VERSION : 0.1
   VAR_INPUT
      IN1 : DInt;
      IN2 : DInt;
      IN3 : DInt;
      IN4 : DInt;
      IN5 : DInt;
      IN6 : DInt;
      IN7 : DInt;
   END_VAR
   VAR_OUTPUT
      Out : Real;
   END_VAR
BEGIN

REGION Network 2 (SCL)
   #Out := (DINT_TO_REAL(#IN1 + #IN2 + #IN3) - DINT_TO_REAL(#IN4 + #IN5 + #IN6)) / #IN7;
END_REGION
END_FUNCTION_BLOCK

FUNCTION_BLOCK "PGC Flush"   // FB517, LAD
{ S7_Optimized_Access := 'TRUE' }
VERSION : 0.1
   VAR_INPUT
      Activate : Bool;
      Override : Bool;
      "PGC Purge Duration" : Time := T#60m;
      "Temperature Setpoint" : Real := 50.0;
      Temperature : Real;
      "PGC Stop Delay" : Time := T#10m;
      "PGC Stoped" : Bool;
      "CAB Started" : Bool;
      "CAB after Start Delay" : Time := T#60s;
      "CAB RPM Cmd" : Real := 400.0;
      "IGG Mode" : Int;   // 1 = Auto, 2 = Man, 3 = FatAuto, 4 = FatMan
      "IGG Stoped" : Bool;
      Alarm : Bool;
      "CV405 Opened" : Real;
      "CV403 Opened" : Real;
      "CV401 Opened" : Bool;
      "CV441 Closed" : Bool;
      "CV431 Opened" : Bool;
   END_VAR
   VAR_OUTPUT
      "CV405 Open" : Bool;
      "CV403 Open" : Bool;
      "CV401 Open" : Bool;
      "CV441 Close" : Bool;
      "CV431 Open" : Bool;
      "CAB Start" : Bool;
      "CAB RPM Ctrl" : Real;
      "CV403 Modulate" : Bool;
      Running : Bool;
      "Stop PGC" : Bool;
      Done : Bool;
   END_VAR
   VAR
      "CAB earlier Stop Aux" : Time;
      "PGC Stop Delay TON" : TON_TIME;
      "Sequence Max Time TON" : TON_TIME;
      "CAB after Start Delay TON" : TON_TIME;
      "Flip Flop_Override" : "Flip Flop";
      "CAB earlier STOP" : TON_TIME;
      "Valve to origin Delay" : TOF_TIME;
      "Valve Opened Delay" : TOF_TIME;
      "PGC Stop Puls" : TP_TIME;
      "Modulate Delay" : TON_TIME;
      "CAB after Start Delay Aux" : Bool;
   END_VAR
BEGIN

REGION Network 1
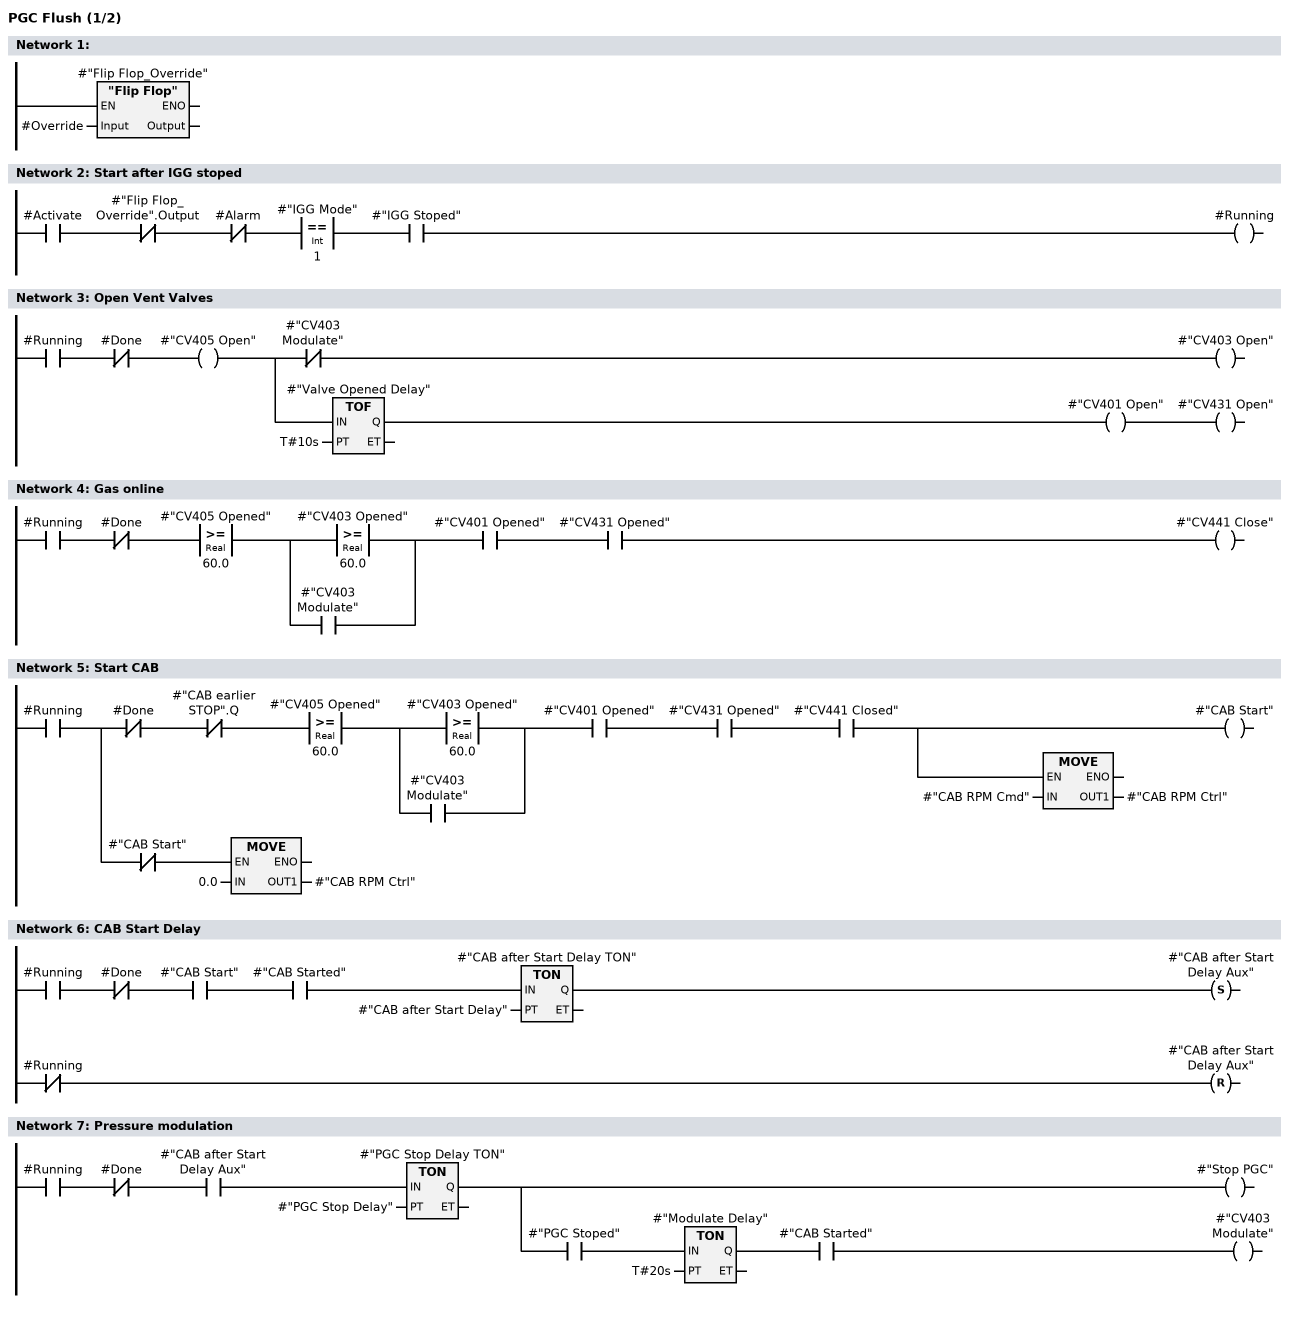
   RUNG wire#powerrail
      #"Flip Flop_Override"(Input := #Override, Output =>)
   END_RUNG
   // the same network as SCL:
   #"Flip Flop_Override"(Input := #Override);   // "Flip Flop"
END_REGION

REGION Network 2: Start after IGG stoped
   RUNG wire#powerrail
      Contact( #Activate )
      I_Contact( #"Flip Flop_Override".Output )
      I_Contact( #Alarm )
      { S7_Templates := "SrcType := Int" } EQ_Contact(in1 := #"IGG Mode", in2 := 1)
      Contact( #"IGG Stoped" )
      Coil( #Running )
   END_RUNG
   // the same network as SCL:
   #Running := #Activate AND NOT #"Flip Flop_Override".Output AND NOT #Alarm AND (#"IGG Mode" = 1) AND #"IGG Stoped";
END_REGION

REGION Network 3: Open Vent Valves
   #"CV405 Open" := #Running AND NOT #Done;
   #"CV403 Open" := #"CV405 Open" AND NOT #"CV403 Modulate";
   #"Valve Opened Delay"(IN := #"CV405 Open", PT := T#10s);   // TOF
   #"CV401 Open" := #"Valve Opened Delay".Q;
   #"CV431 Open" := #"Valve Opened Delay".Q;
END_REGION

REGION Network 4: Gas online
   RUNG wire#powerrail
      Contact( #Running )
      I_Contact( #Done )
      { S7_Templates := "SrcType := Real" } GE_Contact(in1 := #"CV405 Opened", in2 := 60.0)
      wire#w1
      { S7_Templates := "SrcType := Real" } GE_Contact(in1 := #"CV403 Opened", in2 := 60.0)
      wire#w2
      Contact( #"CV401 Opened" )
      Contact( #"CV431 Opened" )
      Coil( #"CV441 Close" )
   END_RUNG
   RUNG wire#w1
      Contact( #"CV403 Modulate" )
   END_RUNG wire#w2
   // the same network as SCL:
   #"CV441 Close" := #Running AND NOT #Done AND (#"CV405 Opened" >= 60.0) AND ((#"CV403 Opened" >= 60.0) OR #"CV403 Modulate") AND #"CV401 Opened" AND #"CV431 Opened";
END_REGION

REGION Network 5: Start CAB
   RUNG wire#powerrail
      Contact( #Running )
      wire#w1
      I_Contact( #Done )
      I_Contact( #"CAB earlier STOP".Q )
      { S7_Templates := "SrcType := Real" } GE_Contact(in1 := #"CV405 Opened", in2 := 60.0)
      wire#w2
      { S7_Templates := "SrcType := Real" } GE_Contact(in1 := #"CV403 Opened", in2 := 60.0)
      wire#w3
      Contact( #"CV401 Opened" )
      Contact( #"CV431 Opened" )
      Contact( #"CV441 Closed" )
      wire#w4
      Coil( #"CAB Start" )
   END_RUNG
   RUNG wire#w2
      Contact( #"CV403 Modulate" )
   END_RUNG wire#w3
   RUNG wire#w4
      Move(in := #"CAB RPM Cmd", out1 => #"CAB RPM Ctrl")
   END_RUNG
   RUNG wire#w1
      I_Contact( #"CAB Start" )
      Move(in := 0.0, out1 => #"CAB RPM Ctrl")
   END_RUNG
   // the same network as SCL:
   #"CAB Start" := #Running AND NOT #Done AND NOT #"CAB earlier STOP".Q AND (#"CV405 Opened" >= 60.0) AND ((#"CV403 Opened" >= 60.0) OR #"CV403 Modulate") AND #"CV401 Opened" AND #"CV431 Opened" AND #"CV441 Closed";
   IF #"CAB Start" THEN #"CAB RPM Ctrl" := #"CAB RPM Cmd"; END_IF;
   IF #Running AND NOT #"CAB Start" THEN #"CAB RPM Ctrl" := 0.0; END_IF;
END_REGION

REGION Network 6: CAB Start Delay
   #"CAB after Start Delay TON"(IN := #Running AND NOT #Done AND #"CAB Start" AND #"CAB Started",   // TON
                           PT := #"CAB after Start Delay");
   IF #"CAB after Start Delay TON".Q THEN #"CAB after Start Delay Aux" := TRUE; END_IF;
   IF NOT #Running THEN #"CAB after Start Delay Aux" := FALSE; END_IF;
END_REGION

REGION Network 7: Pressure modulation
   #"PGC Stop Delay TON"(IN := #Running AND NOT #Done AND #"CAB after Start Delay Aux", PT := #"PGC Stop Delay");   // TON
   #"Stop PGC" := #"PGC Stop Delay TON".Q;
   #"Modulate Delay"(IN := #"PGC Stop Delay TON".Q AND #"PGC Stoped", PT := T#20s);   // TON
   #"CV403 Modulate" := #"Modulate Delay".Q AND #"CAB Started";
END_REGION

REGION Network 8: Sequence max time
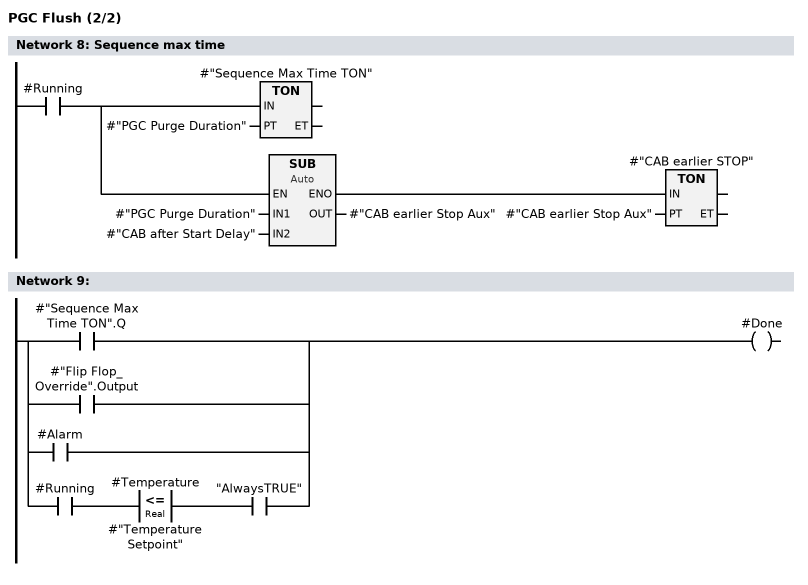
   #"Sequence Max Time TON"(IN := #Running, PT := #"PGC Purge Duration");   // TON
   IF #Running THEN #"CAB earlier Stop Aux" := #"PGC Purge Duration" - #"CAB after Start Delay"; END_IF;
   #"CAB earlier STOP"(IN := #Running, PT := #"CAB earlier Stop Aux");   // TON
END_REGION

REGION Network 9
   RUNG wire#powerrail
      Contact( #"Sequence Max Time TON".Q )
      wire#w1
      Coil( #Done )
   END_RUNG
   RUNG wire#powerrail
      Contact( #"Flip Flop_Override".Output )
   END_RUNG wire#w1
   RUNG wire#powerrail
      Contact( #Alarm )
   END_RUNG wire#w1
   RUNG wire#powerrail
      Contact( #Running )
      { S7_Templates := "SrcType := Real" } LE_Contact(in1 := #Temperature, in2 := #"Temperature Setpoint")
      Contact( "AlwaysTRUE" )
   END_RUNG wire#w1
   // the same network as SCL:
   #Done := #"Sequence Max Time TON".Q OR #"Flip Flop_Override".Output OR #Alarm OR (#Running AND (#Temperature <= #"Temperature Setpoint") AND "AlwaysTRUE");
END_REGION
END_FUNCTION_BLOCK

FUNCTION_BLOCK "RAMP"   // FB518, LAD
{ S7_Optimized_Access := 'TRUE' }
VERSION : 0.1
   VAR_INPUT
      Start : Bool;
      "Time span" : Time;
      "Minimum Value" : Real;
      "Maximum Value" : Real;
   END_VAR
   VAR_OUTPUT
      Value : Real;
      "Ramp Done" : Bool;
   END_VAR
   VAR
      "RUN Time" : TON_TIME;
      "RUN Time Aux" : Real;
      "Time span Aux" : Real;
      "Maximum Value M" : Real;
   END_VAR
BEGIN

REGION Network 1
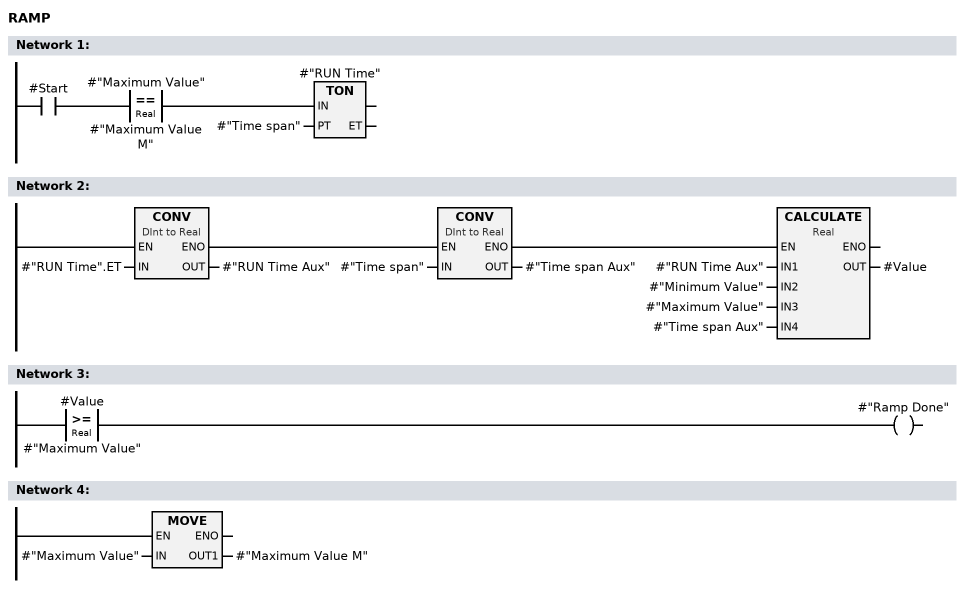
   #"RUN Time"(IN := #Start AND (#"Maximum Value" = #"Maximum Value M"), PT := #"Time span");   // TON
END_REGION

REGION Network 2
   RUNG wire#powerrail
      { S7_Templates := "[SrcType := DInt, DestType := Real]" } Convert(in := #"RUN Time".ET, out => #"RUN Time Aux")
      { S7_Templates := "[SrcType := DInt, DestType := Real]" } Convert(in := #"Time span", out => #"Time span Aux")
      { S7_Templates := "SrcType := Real"; S7_Expression := "((IN1*(IN3-IN2))/IN4)+IN2" } Calculate(in1 := #"RUN Time Aux", in2 := #"Minimum Value", in3 := #"Maximum Value", in4 := #"Time span Aux", out => #Value)
   END_RUNG
   // the same network as SCL:
   #"RUN Time Aux" := DINT_TO_REAL(#"RUN Time".ET);
   #"Time span Aux" := DINT_TO_REAL(#"Time span");
   #Value := ((#"RUN Time Aux"*(#"Maximum Value"-#"Minimum Value"))/#"Time span Aux")+#"Minimum Value";
END_REGION

REGION Network 3
   RUNG wire#powerrail
      { S7_Templates := "SrcType := Real" } GE_Contact(in1 := #Value, in2 := #"Maximum Value")
      Coil( #"Ramp Done" )
   END_RUNG
   // the same network as SCL:
   #"Ramp Done" := #Value >= #"Maximum Value";
END_REGION

REGION Network 4
   RUNG wire#powerrail
      Move(in := #"Maximum Value", out1 => #"Maximum Value M")
   END_RUNG
   // the same network as SCL:
   #"Maximum Value M" := #"Maximum Value";
END_REGION
END_FUNCTION_BLOCK

FUNCTION_BLOCK "Choose Real"   // FB519, LAD
{ S7_Optimized_Access := 'TRUE' }
VERSION : 0.1
   VAR_INPUT
      Choose : Bool;
      "Option 1" : Real;
      "Option 2" : Real;
   END_VAR
   VAR_OUTPUT
      Output : Real;
   END_VAR
   VAR
      True : Bool;
      False : Bool;
      "Option 1 M" : Real;
      "Option 2 M" : Real;
      "Choose Internal" : Bool;
      "Puls Aux" : Struct
         "Puls Aux 1" : Bool;
         "Puls Aux 2" : Bool;
         "Puls Aux 3" : Bool;
         "Puls Aux 4" : Bool;
         "Puls Aux 5" : Bool;
         "Puls Aux 6" : Bool;
      END_STRUCT;
      "TP P CHOOSE1" : TP_TIME;
      "TP N CHOOSE2" : TP_TIME;
      "TP N CHOOSE1" : TP_TIME;
      "TP P CHOOSE2" : TP_TIME;
      R_TRIG_Instance : R_TRIG;
      Puls : TP_TIME;
   END_VAR
   VAR_TEMP   // added for the SCL form of the ladder/FBD networks
      _w1 : Bool;
      _w2 : Bool;
      _w3 : Bool;
      _w4 : Bool;
      _w5 : Bool;
   END_VAR
BEGIN

REGION Network 1: False/True
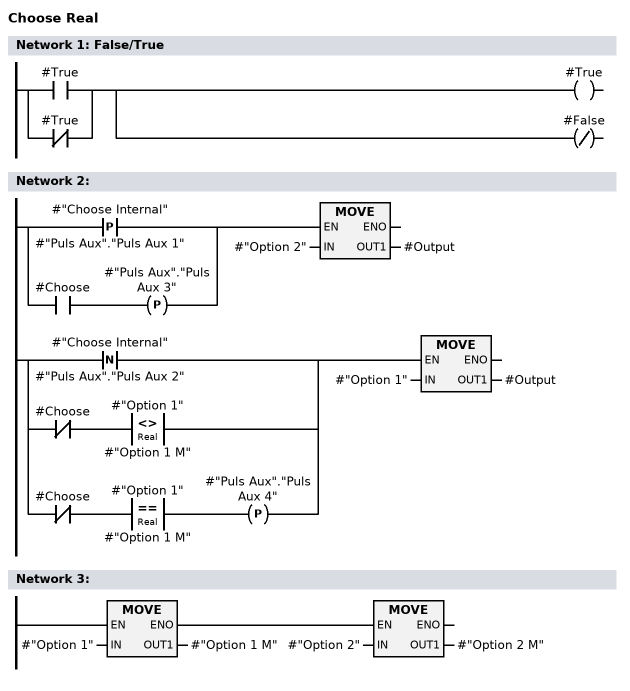
   RUNG wire#powerrail
      Contact( #True )
      wire#w1
      Coil( #True )
   END_RUNG
   RUNG wire#powerrail
      I_Contact( #True )
   END_RUNG wire#w1
   RUNG wire#w1
      I_Coil( #False )
   END_RUNG
   // the same network as SCL:
   #True := #True OR NOT #True;
   #False := NOT #True;
END_REGION

REGION Network 2
   RUNG wire#powerrail
      P_Contact(operand := #"Choose Internal", bit := #"Puls Aux"."Puls Aux 1")
      wire#w1
      Move(in := #"Option 2", out1 => #Output)
   END_RUNG
   RUNG wire#powerrail
      Contact( #Choose )
      P_Trig( #"Puls Aux"."Puls Aux 3" )
   END_RUNG wire#w1
   RUNG wire#powerrail
      N_Contact(operand := #"Choose Internal", bit := #"Puls Aux"."Puls Aux 2")
      wire#w2
      Move(in := #"Option 1", out1 => #Output)
   END_RUNG
   RUNG wire#powerrail
      I_Contact( #Choose )
      { S7_Templates := "SrcType := Real" } NE_Contact(in1 := #"Option 1", in2 := #"Option 1 M")
   END_RUNG wire#w2
   RUNG wire#powerrail
      I_Contact( #Choose )
      { S7_Templates := "SrcType := Real" } EQ_Contact(in1 := #"Option 1", in2 := #"Option 1 M")
      P_Trig( #"Puls Aux"."Puls Aux 4" )
   END_RUNG wire#w2
   // the same network as SCL:
   #_w1 := #"Choose Internal" AND NOT #"Puls Aux"."Puls Aux 1";   // rising edge of #"Choose Internal"
   #"Puls Aux"."Puls Aux 1" := #"Choose Internal";
   #_w2 := #Choose AND NOT #"Puls Aux"."Puls Aux 3";   // rising edge
   #"Puls Aux"."Puls Aux 3" := #Choose;
   IF #_w1 OR #_w2 THEN #Output := #"Option 2"; END_IF;
   #_w3 := NOT #"Choose Internal" AND #"Puls Aux"."Puls Aux 2";   // falling edge of #"Choose Internal"
   #"Puls Aux"."Puls Aux 2" := #"Choose Internal";
   #_w4 := NOT #Choose AND (#"Option 1" = #"Option 1 M");
   #_w5 := #_w4 AND NOT #"Puls Aux"."Puls Aux 4";   // rising edge
   #"Puls Aux"."Puls Aux 4" := #_w4;
   IF #_w3 OR (NOT #Choose AND (#"Option 1" <> #"Option 1 M")) OR #_w5 THEN #Output := #"Option 1"; END_IF;
END_REGION

REGION Network 3
   RUNG wire#powerrail
      Move(in := #"Option 1", out1 => #"Option 1 M")
      Move(in := #"Option 2", out1 => #"Option 2 M")
   END_RUNG
   // the same network as SCL:
   #"Option 1 M" := #"Option 1";
   #"Option 2 M" := #"Option 2";
END_REGION
END_FUNCTION_BLOCK

FUNCTION "Bool to Word" : Void   // FC202, FBD
{ S7_Optimized_Access := 'FALSE' }
VERSION : 0.1
// Die Funktion gruppiert 16 Variablen vom Datentyp "Bool" zu einer Variablen vom Datentyp "Word".
// *******************************************************************************
// The function groups 16 variables with type of data "Bool" to a variable with type of data "Word".
   VAR_INPUT
      Bit0 : Bool;
      Bit1 : Bool;
      Bit2 : Bool;
      Bit3 : Bool;
      Bit4 : Bool;
      Bit5 : Bool;
      Bit6 : Bool;
      Bit7 : Bool;
      Bit8 : Bool;
      Bit9 : Bool;
      Bit10 : Bool;
      Bit11 : Bool;
      Bit12 : Bool;
      Bit13 : Bool;
      Bit14 : Bool;
      Bit15 : Bool;
   END_VAR
   VAR_OUTPUT
      "Word" : Word;
   END_VAR
   VAR_TEMP
      aux : DInt;
   END_VAR
BEGIN

REGION Network 1: aux
   // Setze Hilfsvariable "aux" auf den Anfangswert 0.
   // ***************************************************************************
   // Set the auxiliary variable "aux" to the initial value 0.
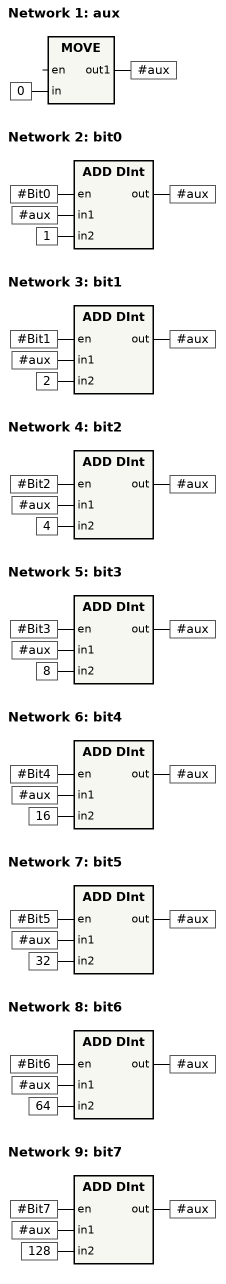
   #aux := 0;
END_REGION

REGION Network 2: bit0
   // Addiere Bit 0 zur Hilfsvariable "aux" vom Datentyp "UInt".
   // ***************************************************************************
   // Add Bit 0 to the auxiliary variable "aux" with type of data "UInt".
   IF #Bit0 THEN #aux := #aux + 1; END_IF;
END_REGION

REGION Network 3: bit1
   // Addiere Bit 1 zur Hilfsvariable "aux".
   // ***************************************************************************
   // Add Bit 1 to the auxiliary variable "aux".
   IF #Bit1 THEN #aux := #aux + 2; END_IF;
END_REGION

REGION Network 4: bit2
   // Addiere Bit 2 zur Hilfsvariable "aux".
   // ***************************************************************************
   // Add Bit 2 to the auxiliary variable "aux".
   IF #Bit2 THEN #aux := #aux + 4; END_IF;
END_REGION

REGION Network 5: bit3
   // Addiere Bit 3 zur Hilfsvariable "aux".
   // ***************************************************************************
   // Add Bit 3 to the auxiliary variable "aux".
   IF #Bit3 THEN #aux := #aux + 8; END_IF;
END_REGION

REGION Network 6: bit4
   // Addiere Bit 4 zur Hilfsvariable "aux".
   // ***************************************************************************
   // Add Bit 4 to the auxiliary variable "aux".
   IF #Bit4 THEN #aux := #aux + 16; END_IF;
END_REGION

REGION Network 7: bit5
   // Addiere Bit 5 zur Hilfsvariable "aux".
   // ***************************************************************************
   // Add Bit 5 to the auxiliary variable "aux".
   IF #Bit5 THEN #aux := #aux + 32; END_IF;
END_REGION

REGION Network 8: bit6
   // Addiere Bit 6 zur Hilfsvariable "aux".
   // ***************************************************************************
   // Add Bit 6 to the auxiliary variable "aux".
   IF #Bit6 THEN #aux := #aux + 64; END_IF;
END_REGION

REGION Network 9: bit7
   // Addiere Bit 7 zur Hilfsvariable "aux".
   // ***************************************************************************
   // Add Bit 7 to the auxiliary variable "aux".
   IF #Bit7 THEN #aux := #aux + 128; END_IF;
END_REGION

REGION Network 10: bit8
   // Addiere Bit 8 zur Hilfsvariable "aux".
   // ***************************************************************************
   // Add Bit 8 to the auxiliary variable "aux".
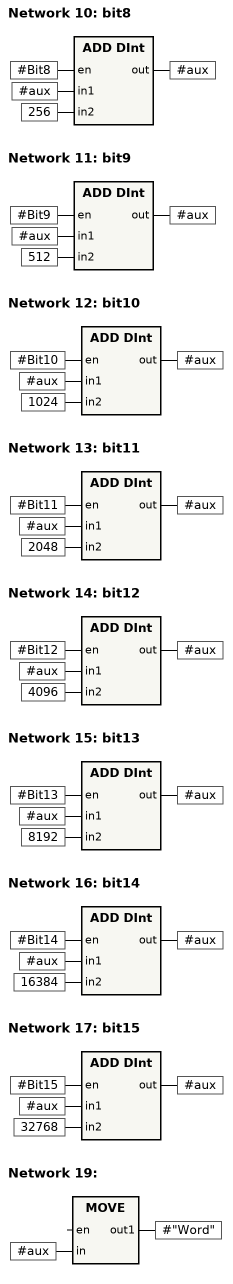
   IF #Bit8 THEN #aux := #aux + 256; END_IF;
END_REGION

REGION Network 11: bit9
   // Addiere Bit 9 zur Hilfsvariable "aux".
   // ***************************************************************************
   // Add Bit 9 to the auxiliary variable "aux".
   IF #Bit9 THEN #aux := #aux + 512; END_IF;
END_REGION

REGION Network 12: bit10
   // Addiere Bit 10 zur Hilfsvariable "aux".
   // ***************************************************************************
   // Add Bit 10 to the auxiliary variable "aux".
   IF #Bit10 THEN #aux := #aux + 1024; END_IF;
END_REGION

REGION Network 13: bit11
   // Addiere Bit 11 zur Hilfsvariable "aux".
   // ***************************************************************************
   // Add Bit 11 to the auxiliary variable "aux".
   IF #Bit11 THEN #aux := #aux + 2048; END_IF;
END_REGION

REGION Network 14: bit12
   // Addiere Bit 12 zur Hilfsvariable "aux".
   // ***************************************************************************
   // Add Bit 12 to the auxiliary variable "aux".
   IF #Bit12 THEN #aux := #aux + 4096; END_IF;
END_REGION

REGION Network 15: bit13
   // Addiere Bit 13 zur Hilfsvariable "aux".
   // ***************************************************************************
   // Add Bit 13 to the auxiliary variable "aux".
   IF #Bit13 THEN #aux := #aux + 8192; END_IF;
END_REGION

REGION Network 16: bit14
   // Addiere Bit 14 zur Hilfsvariable "aux".
   // ***************************************************************************
   // Add Bit 14 to the auxiliary variable "aux".
   IF #Bit14 THEN #aux := #aux + 16384; END_IF;
END_REGION

REGION Network 17: bit15
   // Addiere Bit 15 zur Hilfsvariable "aux".
   // ***************************************************************************
   // Add Bit 15 to the auxiliary variable "aux".
   IF #Bit15 THEN #aux := #aux + 32768; END_IF;
END_REGION

REGION Network 18: Word
   // Der Wert der Variablen "aux" wird  vom Datentyp "UInt" zum Datentyp "Word" konvertiert und der Ausgangsvariablen "Word" übergeben.
   // ***************************************************************************
   // The value of the variable "aux" will convert from type of data "UInt" to type of data "Word" and transfered to the output variable "Word".
END_REGION

REGION Network 19
   #"Word" := #aux;
END_REGION
END_FUNCTION

// folder: 60 - 69 Alarm & Satus Handling

FUNCTION_BLOCK "Tanks Closed"   // FB70, LAD
{ S7_Optimized_Access := 'TRUE' }
VERSION : 0.1
   VAR_INPUT
      "Nr Tanks Activated" : Int;
      Reset : Bool;
   END_VAR
   VAR_OUTPUT
      "Tanks Closed" : Bool;
   END_VAR
   VAR
      R_TRIG_Instance : R_TRIG;
      "NR TANKS ACTIVATED M" : Int;
   END_VAR
BEGIN

REGION Network 1
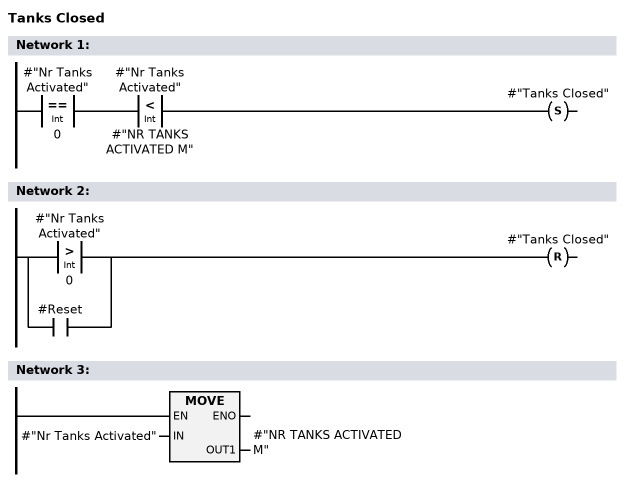
   RUNG wire#powerrail
      { S7_Templates := "SrcType := Int" } EQ_Contact(in1 := #"Nr Tanks Activated", in2 := 0)
      { S7_Templates := "SrcType := Int" } LT_Contact(in1 := #"Nr Tanks Activated", in2 := #"NR TANKS ACTIVATED M")
      S_Coil( #"Tanks Closed" )
   END_RUNG
   // the same network as SCL:
   IF (#"Nr Tanks Activated" = 0) AND (#"Nr Tanks Activated" < #"NR TANKS ACTIVATED M") THEN
       #"Tanks Closed" := TRUE;
   END_IF;
END_REGION

REGION Network 2
   RUNG wire#powerrail
      { S7_Templates := "SrcType := Int" } GT_Contact(in1 := #"Nr Tanks Activated", in2 := 0)
      wire#w1
      R_Coil( #"Tanks Closed" )
   END_RUNG
   RUNG wire#powerrail
      Contact( #Reset )
   END_RUNG wire#w1
   // the same network as SCL:
   IF (#"Nr Tanks Activated" > 0) OR #Reset THEN #"Tanks Closed" := FALSE; END_IF;
END_REGION

REGION Network 3
   RUNG wire#powerrail
      Move(in := #"Nr Tanks Activated", out1 => #"NR TANKS ACTIVATED M")
   END_RUNG
   // the same network as SCL:
   #"NR TANKS ACTIVATED M" := #"Nr Tanks Activated";
END_REGION
END_FUNCTION_BLOCK

FUNCTION "60_Alarms" : Void   // FC60, LAD
TITLE = Alarm Processing
{ S7_Optimized_Access := 'TRUE' }
AUTHOR : JRS
VERSION : 0.1
// To determine alarm conditions
   VAR_TEMP   // added for the SCL form of the ladder/FBD networks
      _w1 : Bool;
   END_VAR
BEGIN

REGION Network 1: DB60 DBX0.0 = BWT Panel E-Stop Pressed
   // GCU_ALARM_WORD_01_BIT_0
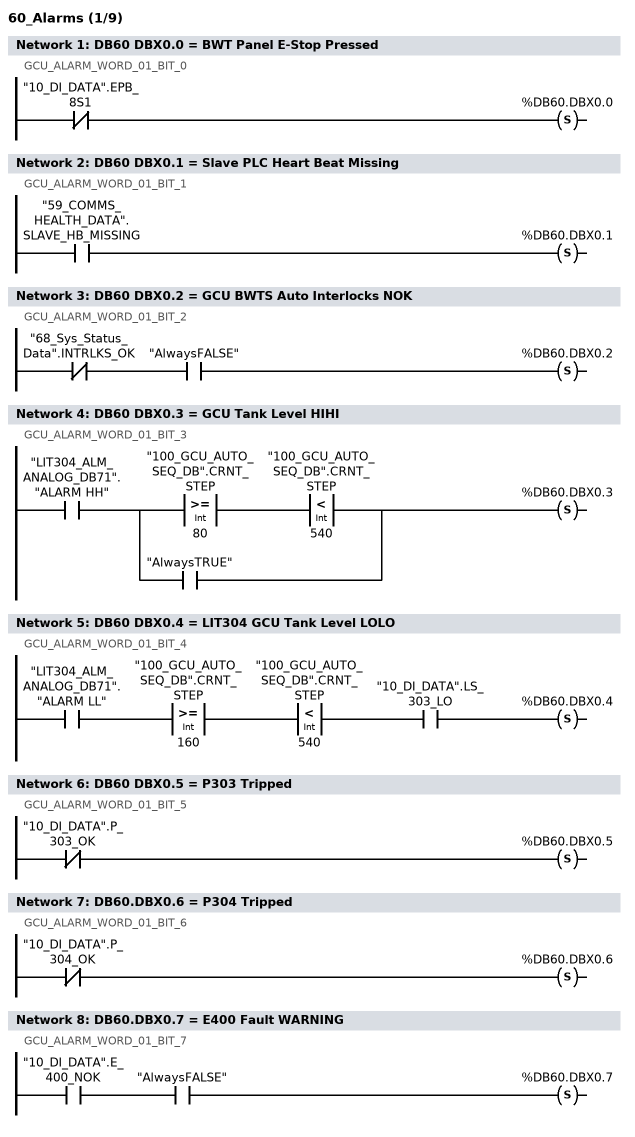
   RUNG wire#powerrail
      I_Contact( "10_DI_DATA".EPB_8S1 )
      S_Coil( %DB60.DBX0.0 )
   END_RUNG
   // the same network as SCL:
   IF NOT "10_DI_DATA".EPB_8S1 THEN %DB60.DBX0.0 := TRUE; END_IF;
END_REGION

REGION Network 2: DB60 DBX0.1 = Slave PLC Heart Beat Missing
   // GCU_ALARM_WORD_01_BIT_1
   RUNG wire#powerrail
      Contact( "59_COMMS_HEALTH_DATA".SLAVE_HB_MISSING )
      S_Coil( %DB60.DBX0.1 )
   END_RUNG
   // the same network as SCL:
   IF "59_COMMS_HEALTH_DATA".SLAVE_HB_MISSING THEN %DB60.DBX0.1 := TRUE; END_IF;
END_REGION

REGION Network 3: DB60 DBX0.2 = GCU BWTS Auto Interlocks NOK
   // GCU_ALARM_WORD_01_BIT_2
   RUNG wire#powerrail
      I_Contact( "68_Sys_Status_Data".INTRLKS_OK )
      Contact( "AlwaysFALSE" )
      S_Coil( %DB60.DBX0.2 )
   END_RUNG
   // the same network as SCL:
   IF NOT "68_Sys_Status_Data".INTRLKS_OK AND "AlwaysFALSE" THEN %DB60.DBX0.2 := TRUE; END_IF;
END_REGION

REGION Network 4: DB60 DBX0.3 = GCU Tank Level HIHI
   // GCU_ALARM_WORD_01_BIT_3
   RUNG wire#powerrail
      Contact( "LIT304_ALM_ANALOG_DB71"."ALARM HH" )
      wire#w1
      { S7_Templates := "SrcType := Int" } GE_Contact(in1 := "100_GCU_AUTO_SEQ_DB".CRNT_STEP, in2 := 80)
      { S7_Templates := "SrcType := Int" } LT_Contact(in1 := "100_GCU_AUTO_SEQ_DB".CRNT_STEP, in2 := 540)
      wire#w2
      S_Coil( %DB60.DBX0.3 )
   END_RUNG
   RUNG wire#w1
      Contact( "AlwaysTRUE" )
   END_RUNG wire#w2
   // the same network as SCL:
   IF "LIT304_ALM_ANALOG_DB71"."ALARM HH" AND ((("100_GCU_AUTO_SEQ_DB".CRNT_STEP >= 80) AND ("100_GCU_AUTO_SEQ_DB".CRNT_STEP < 540)) OR "AlwaysTRUE") THEN
       %DB60.DBX0.3 := TRUE;
   END_IF;
END_REGION

REGION Network 5: DB60 DBX0.4 = LIT304 GCU Tank Level LOLO
   // GCU_ALARM_WORD_01_BIT_4
   RUNG wire#powerrail
      Contact( "LIT304_ALM_ANALOG_DB71"."ALARM LL" )
      { S7_Templates := "SrcType := Int" } GE_Contact(in1 := "100_GCU_AUTO_SEQ_DB".CRNT_STEP, in2 := 160)
      { S7_Templates := "SrcType := Int" } LT_Contact(in1 := "100_GCU_AUTO_SEQ_DB".CRNT_STEP, in2 := 540)
      Contact( "10_DI_DATA".LS_303_LO )
      S_Coil( %DB60.DBX0.4 )
   END_RUNG
   // the same network as SCL:
   IF "LIT304_ALM_ANALOG_DB71"."ALARM LL" AND ("100_GCU_AUTO_SEQ_DB".CRNT_STEP >= 160) AND ("100_GCU_AUTO_SEQ_DB".CRNT_STEP < 540) AND "10_DI_DATA".LS_303_LO THEN
       %DB60.DBX0.4 := TRUE;
   END_IF;
END_REGION

REGION Network 6: DB60 DBX0.5 = P303 Tripped
   // GCU_ALARM_WORD_01_BIT_5
   RUNG wire#powerrail
      I_Contact( "10_DI_DATA".P_303_OK )
      S_Coil( %DB60.DBX0.5 )
   END_RUNG
   // the same network as SCL:
   IF NOT "10_DI_DATA".P_303_OK THEN %DB60.DBX0.5 := TRUE; END_IF;
END_REGION

REGION Network 7: DB60.DBX0.6 = P304 Tripped
   // GCU_ALARM_WORD_01_BIT_6
   RUNG wire#powerrail
      I_Contact( "10_DI_DATA".P_304_OK )
      S_Coil( %DB60.DBX0.6 )
   END_RUNG
   // the same network as SCL:
   IF NOT "10_DI_DATA".P_304_OK THEN %DB60.DBX0.6 := TRUE; END_IF;
END_REGION

REGION Network 8: DB60.DBX0.7 = E400 Fault WARNING
   // GCU_ALARM_WORD_01_BIT_7
   RUNG wire#powerrail
      Contact( "10_DI_DATA".E_400_NOK )
      Contact( "AlwaysFALSE" )
      S_Coil( %DB60.DBX0.7 )
   END_RUNG
   // the same network as SCL:
   IF "10_DI_DATA".E_400_NOK AND "AlwaysFALSE" THEN %DB60.DBX0.7 := TRUE; END_IF;
END_REGION

REGION Network 9: DB60.DBX1.0 = E400 Tripped
   // GCU_ALARM_WORD_01_BIT_8
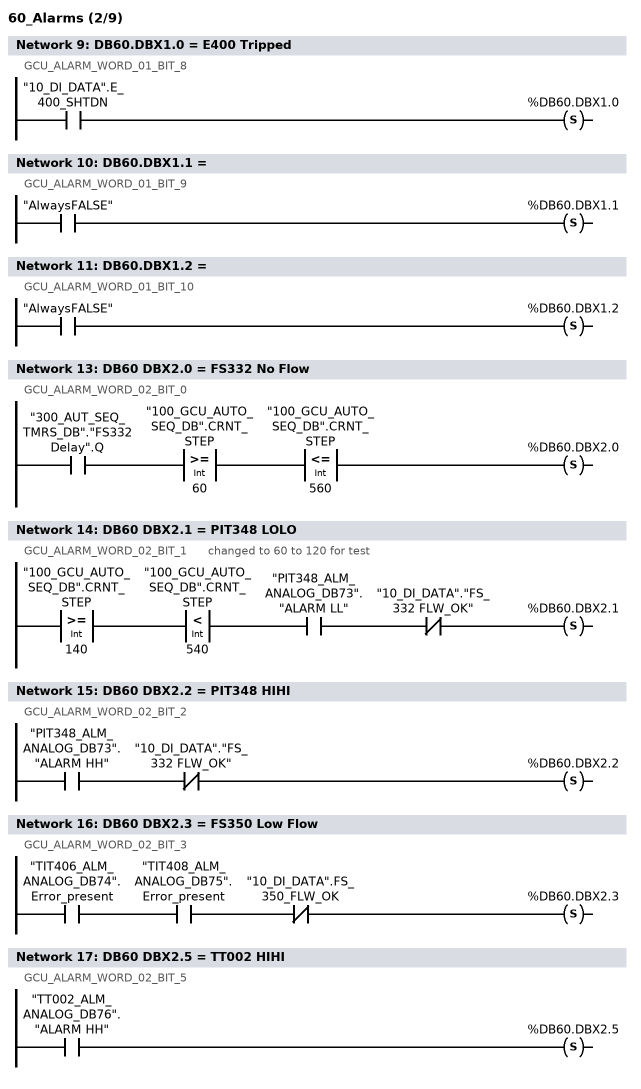
   RUNG wire#powerrail
      Contact( "10_DI_DATA".E_400_SHTDN )
      S_Coil( %DB60.DBX1.0 )
   END_RUNG
   // the same network as SCL:
   IF "10_DI_DATA".E_400_SHTDN THEN %DB60.DBX1.0 := TRUE; END_IF;
END_REGION

REGION Network 10: DB60.DBX1.1 =
   // GCU_ALARM_WORD_01_BIT_9
   RUNG wire#powerrail
      Contact( "AlwaysFALSE" )
      S_Coil( %DB60.DBX1.1 )
   END_RUNG
   // the same network as SCL:
   IF "AlwaysFALSE" THEN %DB60.DBX1.1 := TRUE; END_IF;
END_REGION

REGION Network 11: DB60.DBX1.2 =
   // GCU_ALARM_WORD_01_BIT_10
   RUNG wire#powerrail
      Contact( "AlwaysFALSE" )
      S_Coil( %DB60.DBX1.2 )
   END_RUNG
   // the same network as SCL:
   IF "AlwaysFALSE" THEN %DB60.DBX1.2 := TRUE; END_IF;
END_REGION
